   // ============================================================
   // Returns true if a certain property is set
   // ============================================================
   #LKinLang_CheckProperty := (#properties AND #propertyToCheck) = #propertyToCheck;
END_FUNCTION

FUNCTION "LKinLang_CreateParameterLookUpTable" : Void   // FC35462, SCL
TITLE = LKinLang_CreateParameterLookUpTable
{ S7_Optimized_Access := 'TRUE' }
AUTHOR : tech.team.motioncontrol@siemens.com
FAMILY : LKinLang
VERSION : 1.1
// The FC creates the parameter look up table for later use in parser
   VAR_INPUT
      language : Int;   // language the lookUpTable should be created for
      mode : Bool;   // 0: Commands with ParameterNameNo 1: Commands without ParameterNameNumber
   END_VAR
   VAR_OUTPUT
      error : Bool;   // TRUE: An error occurred during the execution of the FC
      lastIndexLookUp : DInt;   // last index in lookUpTable
   END_VAR
   VAR_IN_OUT
      parameterLookUpTable : Array[1.."LKINLANG_MAX_NUMBER_OF_PARAMETERS"] of "LKinLang_typeParameterLookUp";   // created parameterLookUpTable
      parameterDefaults : Variant;   // parameter defaults
      parameterCounter : Int;   // parameter counter
      errorString : String;   // error information (textual)
   END_VAR
   VAR_TEMP
      tempParameterIndex : Int;
      tempParameterDefinition : "LKinLang_typeParameterDefinition";
      tempCounter : Int;
      tempSeparator : Array[1.."LKINLANG_NUMBER_OF_SEPARATORS"] of Byte;
      tempMerger : Array[1.."LKINLANG_NUMBER_OF_MERGERS"] of Byte;
      tempParameterDefinitionEmpty : "LKinLang_typeParameterDefinition";
      tempFollowValueCounter : Int;
      tempValidCounts : "LKinLang_typePathDataElementCounter";
      tempString : "LKinLang_typeVariableDeclaration";
      tempKeyToken : "LKinLang_typeKeyToken";
   END_VAR
BEGIN
   //==========================================================================================
   // SIEMENS AG
   // (c)Copyright 2019 All Rights Reserved
   //------------------------------------------------------------------------------------------
   // Library: LKinLang
   // Tested with: S7-1517T-3 PN/DP
   // Engineering: TIA Portal V15
   // Restrictions: ---
   // Requirements: S7-1500T FW 2.5
   // Functionality: LKinLang_CreateParameterLookUpTable
   // The FC creates the parameter look up table for later use in parser
   // 
   // Support: tech.team.motioncontrol@siemens.com
   // Note: Parameter comments are only available in language 'English (United States)'
   //------------------------------------------------------------------------------------------
   // Change log table:
   // Version    Date          Expert in charge    Changes applied
   // 01.00.00   28.05.2019    FR                  First created version
   // 01.00.02   29.07.2019    FR                  Mode now part of internal IF condition
   //===========================================================================================


   //======================================================================
   // Is token a known parameter - return: parameter number for array
   //======================================================================
   // Initialize
   #tempCounter := 0;
   #tempParameterIndex := 0;

   // Check for vallid parameters
   WHILE #tempParameterIndex <> -1 DO
     "LKinLang_SelectLangPackage"(language := #language,
                                  variableDeclarations=>#tempString,
                                  keyToken=>#tempKeyToken,
                                  parameterDefinition := #tempParameterDefinition,
                                  separators => #tempSeparator,
                                  mergers => #tempMerger,
                                  validCounts => #tempValidCounts,
                                  parameterNumber := #tempParameterIndex,
                                  parameterDefaults := #parameterDefaults);


     IF (#tempParameterIndex > -1 AND #tempParameterDefinition.parameterNameNumber <> -1 AND #mode = 0) // Check parameters with parameter number (>-1)
       OR (#tempParameterIndex > -1 AND #tempParameterDefinition.parameterNameNumber = -1 AND #mode = 1) // Check parameters without parameter number (=-1)
     THEN
       #parameterLookUpTable[#parameterCounter].parameterNameString := #tempParameterDefinition.parameterNameString;
       #parameterLookUpTable[#parameterCounter].parameterNameNumber := #tempParameterDefinition.parameterNameNumber;
       #parameterLookUpTable[#parameterCounter].parameterNumber := #tempParameterIndex;

       IF #tempParameterDefinition.priorities <> #tempParameterDefinitionEmpty.priorities THEN
         #parameterLookUpTable[#parameterCounter].directValueWord.%X0 := true;
       END_IF;

       IF #tempParameterDefinition.priorities.cmdCoordinates <> #tempParameterDefinitionEmpty.priorities.cmdCoordinates THEN
         #parameterLookUpTable[#parameterCounter].directValueWord.%X1 := true;
       END_IF;

       IF #tempParameterDefinition.priorities.cmdParameters <> #tempParameterDefinitionEmpty.priorities.cmdParameters THEN
         #parameterLookUpTable[#parameterCounter].directValueWord.%X2 := true;
       END_IF;
       IF #tempParameterDefinition.priorities.cmdParameters.pathDynamics <> #tempParameterDefinitionEmpty.priorities.cmdParameters.pathDynamics THEN
         #parameterLookUpTable[#parameterCounter].directValueWord.%X3 := true;
       END_IF;
       IF #tempParameterDefinition.priorities.cmdParameters.circleParameters <> #tempParameterDefinitionEmpty.priorities.cmdParameters.circleParameters THEN
         #parameterLookUpTable[#parameterCounter].directValueWord.%X4 := true;
       END_IF;

       FOR #tempFollowValueCounter := 1 TO "LKINLANG_NUMBER_OF_FOLLOW_VALUES" DO
         IF #tempParameterDefinition.followingValues[#tempFollowValueCounter] <> #tempParameterDefinitionEmpty.followingValues[#tempFollowValueCounter] THEN
           #parameterLookUpTable[#parameterCounter].followValueWords[#tempFollowValueCounter].%X0 := TRUE;
         END_IF;

         IF #tempParameterDefinition.followingValues[#tempFollowValueCounter].cmdCoordinates <> #tempParameterDefinitionEmpty.followingValues[#tempFollowValueCounter].cmdCoordinates THEN
           #parameterLookUpTable[#parameterCounter].followValueWords[#tempFollowValueCounter].%X1 := TRUE;
         END_IF;

         IF #tempParameterDefinition.followingValues[#tempFollowValueCounter].cmdParameters <> #tempParameterDefinitionEmpty.followingValues[#tempFollowValueCounter].cmdParameters THEN
           #parameterLookUpTable[#parameterCounter].followValueWords[#tempFollowValueCounter].%X2 := TRUE;
         END_IF;

         IF #tempParameterDefinition.followingValues[#tempFollowValueCounter].cmdParameters.pathDynamics <> #tempParameterDefinitionEmpty.followingValues[#tempFollowValueCounter].cmdParameters.pathDynamics THEN
           #parameterLookUpTable[#parameterCounter].followValueWords[#tempFollowValueCounter].%X3 := TRUE;
         END_IF;

         IF #tempParameterDefinition.followingValues[#tempFollowValueCounter].cmdParameters.circleParameters <> #tempParameterDefinitionEmpty.followingValues[#tempFollowValueCounter].cmdParameters.circleParameters THEN
           #parameterLookUpTable[#parameterCounter].followValueWords[#tempFollowValueCounter].%X4 := TRUE;
         END_IF;
       END_FOR;

       #parameterCounter += 1;
       #lastIndexLookUp := #parameterCounter;

       // Check ParameterCounter for Overflow
       IF #parameterCounter > "LKINLANG_MAX_NUMBER_OF_PARAMETERS" THEN
         #error := TRUE;
         #errorString := CONCAT(IN1 := #errorString, IN2 := 'Error: Array overflow lookUp table; Increase "LKINLANG_MAX_NUMBER_OF_PARAMETERS"');
         RETURN;
       END_IF;

     ELSE
       ;// no match
     END_IF;

     #tempCounter += 1;

     // Abort searching when tempParameterIndex = -1
     IF #tempParameterIndex <> -1 THEN
       #tempParameterIndex := #tempCounter;
     END_IF;

   END_WHILE;
END_FUNCTION

FUNCTION "LKinLang_DeleteComment" : Void   // FC35463, SCL
TITLE = LKinLang_DeleteComment
{ S7_Optimized_Access := 'TRUE' }
AUTHOR : tech.team.motioncontrol@siemens.com
FAMILY : LKinLang
VERSION : 1.1
// The FC deletes comments from a given string
   VAR_IN_OUT
      codeline : String;   // line to edit by deleting comments
   END_VAR
   VAR_TEMP
      tempPosOfCommentSign : Int;   // temporary variable for position of found comments
   END_VAR
BEGIN
   //==========================================================================================
   // SIEMENS AG
   // (c)Copyright 2019 All Rights Reserved
   //------------------------------------------------------------------------------------------
   // Library: LKinLang
   // Tested with: S7-1517T-3 PN/DP
   // Engineering: TIA Portal V15
   // Restrictions: ---
   // Requirements: S7-1500T FW 2.5
   // Functionality: LKinLang_DeleteComment
   // The FC deletes comments from a given string
   // 
   // Support: tech.team.motioncontrol@siemens.com
   // Note: Parameter comments are only available in language 'English (United States)'
   //------------------------------------------------------------------------------------------
   // Change log table:
   // Version    Date          Expert in charge    Changes applied
   // 01.00.00   28.05.2019    FR                  First created version
   //===========================================================================================

   //======================================================================
   // Delete comment in referenced ascii line
   //======================================================================  

   // Search semicolon
   #tempPosOfCommentSign := FIND(IN1 := #codeline, IN2 := ';');
   // Get line without comment
   IF #tempPosOfCommentSign <> 0 THEN
     #codeline := MID(IN := #codeline, L := #tempPosOfCommentSign - 1, P := 1);
   END_IF;
END_FUNCTION

FUNCTION "LKinLang_DeleteMoreThanOneSpaceInRow" : Void   // FC35464, SCL
TITLE = LKinLang_DeleteMoreThanOneSpaceInRow
{ S7_Optimized_Access := 'TRUE' }
AUTHOR : tech.team.motioncontrol@siemens.com
FAMILY : LKinLang
VERSION : 1.1
// The FC deletes spaces if there are more than one in a row
   VAR_IN_OUT
      codeLine : String;   // line to edit by deleting multiple spaces
   END_VAR
   VAR_TEMP
      tempCodeLine : String["LKINLANG_LENGTH_OF_ASCII_LINE_STRING"];   // temporary variable to store string
      tempSignCounter : Int;   // temporary variable to count signs
      tempSpaceCounter : Int;   // temporary variable to count spaces
      tempStringLength : Int;   // temporary variable to store string length
      tempSpaceIndex : Int;   // temporary variable to store space index
   END_VAR
   VAR CONSTANT
      SPACE : Byte := 16#20;   // space identifier in ascii code
   END_VAR
BEGIN
   //==========================================================================================
   // SIEMENS AG
   // (c)Copyright 2019 All Rights Reserved
   //------------------------------------------------------------------------------------------
   // Library: LKinLang
   // Tested with: S7-1517T-3 PN/DP
   // Engineering: TIA Portal V15
   // Restrictions: ---
   // Requirements: S7-1500T FW 2.5
   // Functionality: LKinLang_DeleteComment
   // The FC deletes spaces if there are more than one in a row
   // 
   // Support: tech.team.motioncontrol@siemens.com
   // Note: Parameter comments are only available in language 'English (United States)'
   //------------------------------------------------------------------------------------------
   // Change log table:
   // Version    Date          Expert in charge    Changes applied
   // 01.00.00   28.05.2019    FR                  First created version
   //===========================================================================================

   //======================================================================
   // Delete more than one spaces
   //====================================================================== 

   // First delete all spaces on start and end
   // -----------------------------------------------------
   // Count spaces on start ---
   #tempSignCounter := 1;

   WHILE #codeLine[#tempSignCounter] = #SPACE DO
     #tempSignCounter := #tempSignCounter + 1;
   END_WHILE;

   // Spaces
   #codeLine := RIGHT(IN := #codeLine,
                      L := LEN(#codeLine) - (#tempSignCounter - 1));


   // Count spaces on end --- 
   #tempSignCounter := LEN(#codeLine);
   WHILE #codeLine[#tempSignCounter] = #SPACE DO
     #tempSpaceCounter := #tempSpaceCounter + 1;
     #tempSignCounter := #tempSignCounter - 1;
   END_WHILE;

   #codeLine := LEFT(IN := #codeLine,
                     L := LEN(#codeLine) - #tempSpaceCounter);
   #tempSpaceCounter := 0;
   // -----------------------------------------------------

   (* // Too slow FR 2019.03.13
   // Delete more than one space in the middle
   // Testing new approach FR
   // 
   #tempSpaceIndex := FIND(IN1 := #codeLine, IN2 := '  ');

   WHILE #tempSpaceIndex <> 0 DO
     #codeLine := DELETE(IN := #codeLine, L := 1, P := #tempSpaceIndex);
     #tempSpaceIndex := FIND(IN1 := #codeLine, IN2 := '  ');
   END_WHILE;

   #codeLine := #codeLine;*)


    // Check if double space is somewhere in the codeline FR 2019.03.12
   IF FIND(IN1 := #codeLine, IN2 := '  ') <> 0 THEN
     // Delete more than one space in the middle
     #tempStringLength := LEN(#codeLine);

     FOR #tempSignCounter := 1 TO (#tempStringLength) DO
       // First character
       IF #tempSignCounter = 1 AND
         #codeLine[#tempSignCounter] <> #SPACE
       THEN
         #tempCodeLine[#tempSignCounter] := #codeLine[#tempSignCounter];

         // Last character                
       ELSIF #tempSignCounter = #tempStringLength AND
         #codeLine[#tempSignCounter] <> #SPACE
       THEN
         #tempCodeLine[#tempSignCounter - #tempSpaceCounter] := #codeLine[#tempSignCounter];

         // Between first and last character
       ELSIF #tempSignCounter > 1 AND #tempSignCounter < #tempStringLength
       THEN
         // More than one spaces in a row?
         IF #codeLine[#tempSignCounter] = #SPACE AND #codeLine[#tempSignCounter + 1] = #SPACE
         THEN
           // Increment space counter
           #tempSpaceCounter := #tempSpaceCounter + 1;
         ELSE
           // Only one Space
           #tempCodeLine[#tempSignCounter - #tempSpaceCounter] := #codeLine[#tempSignCounter];
         END_IF;

         // Increment space counter if the first or last character is a space 
       ELSE
         #tempSpaceCounter := #tempSpaceCounter + 1;
       END_IF;
     END_FOR;

     // set processed code line to in_out parameter
     #codeLine := #tempCodeLine;

   ELSE
     ;// Do nothing - already finished
     //#codeLine := #codeLine;
   END_IF;
END_FUNCTION

FUNCTION "LKinLang_IsTokenMath" : Bool   // FC35465, SCL
TITLE = LKinLang_IsTokenMath
{ S7_Optimized_Access := 'TRUE' }
AUTHOR : tech.team.motioncontrol@siemens.com
FAMILY : LKinLang
VERSION : 1.1
// Checks if a token is a math expression
   VAR_INPUT
      token : String;   // Token to check
   END_VAR
   // Ret_Val : TRUE: Token is math expression; FALSE: Token is not a math expression
BEGIN
   //==========================================================================================
   // SIEMENS AG
   // (c)Copyright 2019 All Rights Reserved
   //------------------------------------------------------------------------------------------
   // Library: LKinLang
   // Tested with: S7-1517T-3 PN/DP
   // Engineering: TIA Portal V15
   // Restrictions: ---
   // Requirements: S7-1500T FW 2.5
   // Functionality: LKinLang_IsTokenMath
   // The FC checks if a given token is a math expression
   // 
   // Support: tech.team.motioncontrol@siemens.com
   // Note: Parameter comments are only available in language 'English (United States)'
   //------------------------------------------------------------------------------------------
   // Change log table:
   // Version    Date          Expert in charge    Changes applied
   // 01.00.00   17.07.2019    FR                  First created version
   //===========================================================================================

   // Check if token is a valid math expression
   IF #token = 'SIN'
     OR #token = 'COS'  
     OR #token = 'SQR'
     OR #token = 'SQRT'
     OR #token = 'sin'
     OR #token = 'cos'
     OR #token = 'sqr'
     OR #token = 'sqrt'
   THEN
     #LKinLang_IsTokenMath := TRUE; // return true if regular math expression
   ELSE
     #LKinLang_IsTokenMath := FALSE; // return false if not
   END_IF;
END_FUNCTION

FUNCTION "LKinLang_GetValue" : DWord   // FC35466, SCL
TITLE = LKinLang_GetValue
{ S7_Optimized_Access := 'TRUE' }
AUTHOR : tech.team.motioncontrol@siemens.com
FAMILY : LKinLang
VERSION : 1.1
// The FC gets the numerical value of a given string expression
   VAR_INPUT
      tokenNo : Int;   // token number to get the numerical value for
      properties : DWord;   // properties to be considered
      followValCounter : Int;   // counter for follow value
   END_VAR
   VAR_OUTPUT
      parameterValue : LReal;   // numerical value of the expression
   END_VAR
   VAR_IN_OUT
      stringExpression : String;   // string to be checked
      errorString : String;   // error information (textual)
      token : "LKinLang_typeLineTokens";   // token information
   END_VAR
   VAR_TEMP
      tempSeparatorFound : Bool;   // temporary variable for found / not found separator
      tempStringExpression : String;   // temporary variable for storage of string expression
      tempStringLength : Int;   // temporary variable for string length
      tempCounter : Int;   // temporary counter variable
      tempSeparatorCounter : Int;   // temporary counter variable for separators
      tempTokenOffset : Int;   // temporary variable for offset of token
      tempMathParserResult : Struct   // temporary variable for math parser result
         finalResult : LReal;
         errorID : DInt;
      END_STRUCT;
   END_VAR
   VAR CONSTANT
      REAL_MIN : LReal := -3.402823E+38;
      REAL_MAX : LReal := 3.402823E+38;
      DINT_MIN : DInt := -2147483648;
      DINT_MAX : DInt := +2147483647;
      INT_MIN : Int := -32768;
      INT_MAX : Int := 32767;
      ERR_PARAMETER_COUNTER : DWord := 16#8001;
      ERR_SYNTAX_MATH_EXPRESSION : DWord := 16#8002;
      ERR_SYNTAX_PARAMETER : DWord := 16#8003;
      ERR_PARAMETER_OVERFLOW : DWord := 16#8004;
      ERR_ALREADY_SET : DWord := 16#8005;
      WARN_NO_MORE_VALUES : DWord := 16#7100;
      COMMA : Char := ',';
   END_VAR
BEGIN
   //==========================================================================================
   // SIEMENS AG
   // (c)Copyright 2019 All Rights Reserved
   //------------------------------------------------------------------------------------------
   // Library: LKinLang
   // Tested with: S7-1517T-3 PN/DP
   // Engineering: TIA Portal V15
   // Restrictions: ---
   // Requirements: S7-1500T FW 2.5
   // Functionality: LKinLang_GetValue
   // The FC gets the numerical value of a given string expression
   // 
   // Support: tech.team.motioncontrol@siemens.com
   // Note: Parameter comments are only available in language 'English (United States)'
   //------------------------------------------------------------------------------------------
   // Change log table:
   // Version    Date          Expert in charge    Changes applied
   // 01.00.00   28.05.2019    FR                  First created version
   // 01.00.01   16.01.2020    FR                  Updated to work with H functions
   //===========================================================================================

   // Initialize variables
   #LKinLang_GetValue := 0;
   #parameterValue := 0;

   // Check if the string expression contains a function separator (COMMA in this case)
   // If true copy only the string expression until the separator and leave the rest (and delete the first separator)
   #tempStringLength := LEN(#stringExpression);

   // Check for comma in stringExpression
   FOR #tempCounter := 1 TO #tempStringLength DO
     // Search for separator 
     IF #stringExpression[#tempCounter] = #COMMA THEN
       #tempSeparatorFound := TRUE;
       EXIT;
     ELSE
       #tempSeparatorFound := FALSE;
     END_IF;
   END_FOR;

   // Check if comma was found
   IF #tempSeparatorFound THEN
     // Copy first value to TempStringExpression 
     #tempStringExpression := LEFT(IN := #stringExpression, L := #tempCounter - 1);
     // Delete first from stringExpression
     #stringExpression := RIGHT(IN := #stringExpression, L := #tempStringLength - #tempCounter);
   ELSE
     #tempStringExpression := #stringExpression;
     #stringExpression := '';
   END_IF;

   IF #tempStringExpression = '' THEN
     // Empty String --> no more Values follow
     // #Lxxx_GetValue := #ERR_SYNTAX_PARAMETER;
     // #errorString := CONCAT(IN1 := #errorString, IN2 := ';Error: Missing assignment'); // Line number is added outside
     // #errorString := CONCAT(IN1 := #errorString, IN2 := INT_TO_STRING(#followValCounter)); // Line number is added outside
     RETURN;
   ELSIF #tempStringExpression = '*' THEN
     // Do not set this value
     RETURN;
   END_IF;

   IF #followValCounter > 1 THEN
     #tempSeparatorCounter := 1;
     // Check for line token offset
     FOR #tempCounter := #tokenNo TO 1 BY -1 DO
       IF #token.lineToken[#tempCounter] = #COMMA OR #token.lineToken[#tempCounter]= '=' THEN
         #tempSeparatorCounter += 1;
       END_IF;

       IF #tempSeparatorCounter = #followValCounter THEN
         EXIT;
       END_IF;
     END_FOR;
     #tempTokenOffset := #tokenNo - #tempCounter;
   ELSE
     #tempCounter := 0;
     #tempTokenOffset := 0;
   END_IF;

   // Calc LReal value --> Check Equation
   REGION GET_VALUE
     IF "LKinLang_CheckProperty"(properties := #properties, propertyToCheck := "LKINLANG_EQUATION") THEN
       REGION EQUATION
         // Equation is possible
         // 
         // Check for correct syntax
         // Two possibilities:
         // 1. Only a number after Parameter 
         // --> Equal sign is optional 
         //  --> When no equal sign then no spaces are allowed --> Example: X12
         //  --> When equal sign then one space allowed --> Example: X = 12
         // 2. Expression after Parameter
         // --> Equal sign is mandatory
         //  --> No spaces --> Example: X=12+34
         //  --> One space allowed --> Example: X = 12+34
         // 
         IF "LKinLang_PostEqualsSignWhenExpressionMandCnd"(currentTokenNo := #tokenNo,
                                                             stringExpression := #tempStringExpression,
                                                             tokenOffset := #tempTokenOffset,
                                                             lineToken := #token) 
         THEN
           // Number: just convert string to real
           IF "LKinLang_IsTokenNumberInclSign"(#tempStringExpression) THEN
             // Set parameter
             #parameterValue := STRING_TO_LREAL(#tempStringExpression);
           ELSE
             //FR not necessary //#errorString := CONCAT(IN1 := #errorString, IN2 := CONCAT(IN1 := ';Error: str=', IN2 := #tempStringExpression));
             #tempMathParserResult := "LKinLang_CalcMathAndBool"(inputString := #tempStringExpression);

             // Error with math parser
             //******************************************
             IF #tempMathParserResult.errorID <> 0 THEN
               #LKinLang_GetValue := #ERR_SYNTAX_MATH_EXPRESSION;

               #errorString := CONCAT(IN1 := #errorString, IN2 := CONCAT(IN1 := ';Error: Mathresult=', IN2 := "LKinLang_LRealToReducedString"(input:=#tempMathParserResult.finalResult,decimalPlaces:=4)));
               #errorString := CONCAT(IN1 := #errorString, IN2 := CONCAT(IN1 := ';Error: No=', IN2 := DINT_TO_STRING(#tempMathParserResult.errorID)));
               // Line number is added outside
               //#errorString := CONCAT(IN1 := #errorString, IN2 := DINT_TO_STRING(#token.lineNo));
               RETURN;
               // Math parser delivers a valid result
               //******************************************
             ELSE
               // Set parameter
               #parameterValue := #tempMathParserResult.finalResult;
             END_IF;
           END_IF;
           #tempStringExpression := '';
         ELSE
           // SyntaxError: not "Y =" or "Y19"
           #LKinLang_GetValue := #ERR_SYNTAX_PARAMETER;
           #errorString := CONCAT(IN1 := #errorString, IN2 := ';Error: Incorrect assignment (Y= or Y1)'); // Line number is added outside
           RETURN;
         END_IF;
       END_REGION EQUATION

     ELSE

       REGION NO_EQUATION
         // Equation is not possible
         IF "LKinLang_PostNumberMandCnd"(algebraicSignAllowed := True, currentTokenNo := #tokenNo, tokenOffset := #tempTokenOffset, lineTokens := #token)
         THEN
           IF "LKinLang_IsTokenNumber"(#tempStringExpression) THEN
             IF #followValCounter = 1 THEN
               #parameterValue := STRING_TO_LREAL(#token.lineToken[#tokenNo - 1]);
             ELSE
               #parameterValue := STRING_TO_LREAL(#token.lineToken[#tokenNo - #tempTokenOffset - 1]);
             END_IF;

             // Check if Mxx stands alone, also there could be something like this Mxx=29
             IF STRING_TO_LREAL(#tempStringExpression) = #parameterValue THEN
               #tempStringExpression := '';
             ELSE
               #LKinLang_GetValue := #ERR_SYNTAX_PARAMETER;
               #errorString := CONCAT(IN1 := #errorString, IN2 := ';Error: Incorrect assignment '); // Line number is added outside
               #errorString := CONCAT(IN1 := #errorString, IN2 := INT_TO_STRING(#followValCounter)); // Line number is added outside
               RETURN;
             END_IF;

           ELSIF "LKinLang_IsTokenNumberInclSign"(#tempStringExpression) THEN

             IF #followValCounter = 1 THEN
               #parameterValue := STRING_TO_LREAL(CONCAT(IN1 := #token.lineToken[#tokenNo - 1], IN2 := #token.lineToken[#tokenNo - 2]));
             ELSE
               #parameterValue := STRING_TO_LREAL(CONCAT(IN1 := #token.lineToken[#tokenNo - #tempTokenOffset - 1], IN2 := #token.lineToken[#tokenNo - #tempTokenOffset - 2]));
             END_IF;

             // Check if Mxx stands alone, also there could be something like this Mxx=29
             IF STRING_TO_LREAL(#tempStringExpression) = #parameterValue THEN
               #tempStringExpression := '';
             ELSE
               #LKinLang_GetValue := #ERR_SYNTAX_PARAMETER;
               #errorString := CONCAT(IN1 := #errorString, IN2 := ';Error: Incorrect assignment '); // Line number is added outside
               #errorString := CONCAT(IN1 := #errorString, IN2 := INT_TO_STRING(#followValCounter)); // Line number is added outside
               RETURN;
             END_IF;
           END_IF;
         ELSE
           // SyntaxError: no number after parameter
           #LKinLang_GetValue := #ERR_SYNTAX_PARAMETER;
           #errorString := CONCAT(IN1 := #errorString, IN2 := ';Error: No number after parameter'); // Line number is added outside
           RETURN;
         END_IF;
       END_REGION NO_EQUATION

     END_IF;

   END_REGION GET_VALUE
END_FUNCTION

FUNCTION "LKinLang_EvaluateCondition" : Bool   // FC35467, SCL
TITLE = LKinLang_EvaluateCondition
{ S7_Optimized_Access := 'TRUE' }
AUTHOR : tech.team.motioncontrol@siemens.com
FAMILY : LKinLang
VERSION : 1.0
// Evaluate a given condition for conditional jumps etc.
   VAR_INPUT
      offsetLastTokenIndex : UInt;   // Number of token to skip from end
   END_VAR
   VAR_IN_OUT
      tokenizedLine : "LKinLang_typeLineTokens";   // Actual tokenized line
      varRefList : "LKinLang_typeVarRefList";   // Variables reference list
      localVariables : "LKinLang_typeLocalVariables";   // Local variables array
      interfaceVariables : "LKinLang_typeInterfaceVariables";   // Interface varaibles array
      keyToken : "LKinLang_typeKeyToken";   // Key token to find variables
      subPrgList : "LKinLang_typeSubPrgList";
      errorString : String;   // error string connection
   END_VAR
   VAR_TEMP
      tempStateIntern : Int;   // Internal state
      tempTokenCounter : Int;   // Temporary counter for token
      tempVarType : Int;   // Variable type
      tempVarIndex : Int;   // Variable index in reference list
      tempStringExpression : String;   // Stringexpression
      tempTokenCheck : Struct   // Struct with the token to check / Static struct with the token to check
         actual : String;
         previous : String;
      END_STRUCT;
      tempMathParserResult : "LKinLang_typeMathParserResult";   // Result of math and bool calculation
   END_VAR
   // Ret_Val : Returns result of condition
   VAR CONSTANT
      STATE_IS_TOKEN_VARIABLE : Int := 250;   // Internal FB state: Is token variable
      STATE_TOKEN_IS_VARIABLE : Int := 260;   // Internal FB state: Token is variable
      STATE_TOKEN_IS_UNKNOWN : Int := 270;   // Internal FB state: Token is unknown
      STATE_ERROR : Int := 900;   // Internal FB state: Error
   END_VAR
BEGIN
   //==========================================================================================
   // SIEMENS AG
   // (c)Copyright 2020 All Rights Reserved
   //------------------------------------------------------------------------------------------
   // Library: LKinLang
   // Tested with: S7-1517T-3 PN/DP
   // Engineering: TIA Portal V15
   // Restrictions: ---
   // Requirements: S7-1500T FW 2.5
   // Functionality: LKinLang_EvaluateCondition
   // The FC creates a valid expression for MathParser and returns the result of the calculation
   // 
   // Support: tech.team.motioncontrol@siemens.com
   // Note: Parameter comments are only available in language 'English (United States)'
   //------------------------------------------------------------------------------------------
   // Change log table:
   // Version    Date          Expert in charge    Changes applied
   // 01.00.00   09.01.2019    FR                  First created version
   // 01.00.01   24.11.2020    FR                  Use functions to check if token is a variable
   //===========================================================================================
   //
   // Add everything except " " to the string expression 
   // If it is a variable then replace with the value of the variable
   // Call MathParser to get result of condition

   // There is no left side of equation as the "=" in a condition is not used as a assignment

   // Iterate over all token
   FOR #tempTokenCounter := 1 TO #tokenizedLine.numberOfToken - #offsetLastTokenIndex DO

     // Init variables for each loop
     #tempTokenCheck.actual := #tokenizedLine.lineToken[#tempTokenCounter];

     //Get previous token
     IF #tempTokenCounter > 1 THEN
       #tempTokenCheck.previous := #tokenizedLine.lineToken[#tempTokenCounter - 1];
     ELSE
       #tempTokenCheck.previous := '';
     END_IF;

     // Next state: IS_TOKEN_VARIABLE
     #tempStateIntern := #STATE_IS_TOKEN_VARIABLE;

     // ------------------------------------------------------------------------------------------
     // Is token variable
     // Check if token is a defined variable or interface variable
     // YES: Go to TOKEN_IS_VARIABLE
     // NO: Go to TOKEN_IS_UNKNOWN
     // ------------------------------------------------------------------------------------------ 
     REGION IS_TOKEN_VARIABLE
       IF #tempStateIntern = #STATE_IS_TOKEN_VARIABLE THEN
         // Check if token is a local or interface variable 
         "LKinLang_IsTokenVariable"(lineNumber := #tokenizedLine.lineNo,
                                    tokenCheck := #tempTokenCheck,
                                    varIndex => #tempVarIndex,
                                    varType => #tempVarType,
                                    varRefList := #varRefList,
                                    keyToken := #keyToken,
                                    subPrgList:=#subPrgList,
                                    errorString := #errorString,
                                    stringExpression := #tempStringExpression);

         // Decide where to go next
         IF #errorString <> '' THEN
           // Error occured
           #tempStateIntern := #STATE_ERROR;
           EXIT;
         ELSIF #tempVarIndex <> 0 OR #tempVarType <> 0 THEN
           // Go to "TOKEN_IS_VARIABLE"
           #tempStateIntern := #STATE_TOKEN_IS_VARIABLE;
         ELSE
           // Go to "TOKEN_IS_UNKNOWN"
           #tempStateIntern := #STATE_TOKEN_IS_UNKNOWN;
         END_IF;
       END_IF;
     END_REGION IS_TOKEN_VARIABLE

     // ------------------------------------------------------------------------------------------
     // Token is a variable
     // Token was found to be a valid variable
     // SET or GET value of variable depending on context
     // ------------------------------------------------------------------------------------------ 
     REGION TOKEN_IS_VARIABLE
       IF #tempStateIntern = #STATE_TOKEN_IS_VARIABLE THEN
         // Token is variable 
         // Decide if value of variable has to be set or value must be read
         "LKinLang_GetVariable"(varIndex:=#tempVarIndex,
                                varType:=#tempVarType,
                                localVariables:=#localVariables,
                                interfaceVariables:=#interfaceVariables,
                                stringExpression:=#tempStringExpression);
       END_IF;
     END_REGION TOKEN_IS_VARIABLE

     // ------------------------------------------------------------------------------------------
     // Token is unknown
     // Token is not a parameter or a separator 
     // Check if equation is active and add token to string expression 
     // If token consists of letters, it is a unknown parameter and a error is thrown
     // Always go to TOKEN_PROCESSED
     // ------------------------------------------------------------------------------------------ 
     REGION TOKEN_IS_UNKNOWN
       IF #tempStateIntern = #STATE_TOKEN_IS_UNKNOWN
       THEN
         // Check if actual token is not space --> Copy to StringExpression (e.g. math expressions)
         IF #tempTokenCheck.actual = 'TRUE' THEN
           #tempStringExpression := CONCAT(IN1 := '1', IN2 := #tempStringExpression);
         ELSIF #tempTokenCheck.actual = 'FALSE' THEN
           #tempStringExpression := CONCAT(IN1 := '0', IN2 := #tempStringExpression);
         ELSIF  #tempTokenCheck.actual <> ' ' THEN
           #tempStringExpression := CONCAT(IN1 := #tempTokenCheck.actual, IN2 := #tempStringExpression);
         ELSE
           ; // Do not copy "space"  into string expression
         END_IF;
       END_IF;
     END_REGION TOKEN_IS_UNKNOWN
   END_FOR;

   #LKinLang_EvaluateCondition := FALSE;

   IF #tempStateIntern <> #STATE_ERROR THEN
     // All token are processed 
     // Call MathParser and calculate result
     #tempMathParserResult := "LKinLang_CalcMathAndBool"(inputString := #tempStringExpression);

     // Check for error in math parser
     IF #tempMathParserResult.errorID <> 0
       OR #tempMathParserResult.finalResult < 0
       OR #tempMathParserResult.finalResult > 1
     THEN
       #tempStateIntern := #STATE_ERROR;
       #errorString := CONCAT(IN1 := #errorString, IN2 := ';Error: Cannot evaluate condition ');
       #errorString := CONCAT(IN1 := #errorString, IN2 := #tempStringExpression);
       #errorString := CONCAT(IN1 := #errorString, IN2 := '; in line: ');
       #errorString := CONCAT(IN1 := #errorString, IN2 := UDINT_TO_STRING(#tokenizedLine.lineNo));
     ELSE
       // Math parser delivers a valid result
       // Assign result to value
       #LKinLang_EvaluateCondition := (#tempMathParserResult.finalResult = 1); // If result = 1 then true else false
     END_IF;
   ELSE
     ; // Error occured --> Do nothing
   END_IF;
END_FUNCTION

FUNCTION "LKinLang_IsNewCommand" : Bool   // FC35469, SCL
TITLE = LKinLang_IsNewCommand
{ S7_Optimized_Access := 'TRUE' }
AUTHOR : tech.team.motioncontrol@siemens.com
FAMILY : LKinLang
VERSION : 1.1
// This function checks if a parsed line results in a new PathData command
   VAR_IN_OUT
      actualPathData : "LKinLang_typePathDataElement";   // actual PathData element to be checked
      emptyPathData : "LKinLang_typePathDataElement";   // empty PathData element for comparison
      positioningMode : Int;   // mode for positioning
   END_VAR
   VAR_TEMP
      tempCircMode0 : Bool;   // temporary variable for circMode 0
      tempCircMode1 : Bool;   // temporary variable for circMode 1
      tempCircMode2 : Bool;   // temporary variable for circMode 2
   END_VAR
BEGIN
   //==========================================================================================
   // SIEMENS AG
   // (c)Copyright 2019 All Rights Reserved
   //------------------------------------------------------------------------------------------
   // Library: LKinLang
   // Tested with: S7-1517T-3 PN/DP
   // Engineering: TIA Portal V15
   // Restrictions: ---
   // Requirements: S7-1500T FW 2.5
   // Functionality: LKinLang_IsNewCommand
   // This function checks if a parsed line results in a new PathData command
   // 
   // Support: tech.team.motioncontrol@siemens.com
   // Note: Parameter comments are only available in language 'English (United States)'
   //------------------------------------------------------------------------------------------
   // Change log table:
   // Version    Date          Expert in charge    Changes applied
   // 01.00.00   28.05.2019    FR                  First created version
   // 01.00.01   10.12.2020    FR                  Added case for cmdType=-1
   //===========================================================================================

   #LKinLang_IsNewCommand := 0;

   CASE #actualPathData.pathDataElement.cmdType OF
       -1: // Only check position
           #LKinLang_IsNewCommand := (#actualPathData.priority.cmdCoordinates.cartesianPosition.x > "LKINLANG_PRIO_UNRELEVANT")
           OR (#actualPathData.priority.cmdCoordinates.cartesianPosition.y > "LKINLANG_PRIO_UNRELEVANT")
           OR (#actualPathData.priority.cmdCoordinates.cartesianPosition.z > "LKINLANG_PRIO_UNRELEVANT")
           OR (#actualPathData.priority.cmdCoordinates.cartesianPosition.a > "LKINLANG_PRIO_UNRELEVANT");


     1,2:  // Linear command
       IF #positioningMode = 1 THEN
         // Is it a new absolute position ?
         // Check if last position is same as actual ? --> Do not check could be usefull with flags on same position
         // (#actualPathData.pathDataElement.cmdCoordinates <> #oldPathData.pathDataElement.cmdCoordinates)
         // AND
         //#LKinLang_IsNewCommand := (#actualPathData.pathDataElement.cmdCoordinates.cartesianPosition <> #emptyPathData.pathDataElement.cmdCoordinates.cartesianPosition);
         #LKinLang_IsNewCommand := (#actualPathData.priority.cmdCoordinates.cartesianPosition.x > "LKINLANG_PRIO_UNRELEVANT")
         OR (#actualPathData.priority.cmdCoordinates.cartesianPosition.y > "LKINLANG_PRIO_UNRELEVANT")
         OR (#actualPathData.priority.cmdCoordinates.cartesianPosition.z > "LKINLANG_PRIO_UNRELEVANT")
         OR (#actualPathData.priority.cmdCoordinates.cartesianPosition.a > "LKINLANG_PRIO_UNRELEVANT");

       ELSIF #positioningMode = 2 THEN
         // Is it a new relative position ?
         //#LKinLang_IsNewCommand := (#actualPathData.pathDataElement.cmdCoordinates.cartesianPosition <> #emptyPathData.pathDataElement.cmdCoordinates.cartesianPosition);
         #LKinLang_IsNewCommand := (#actualPathData.priority.cmdCoordinates.cartesianPosition.x > "LKINLANG_PRIO_UNRELEVANT")
         OR (#actualPathData.priority.cmdCoordinates.cartesianPosition.y > "LKINLANG_PRIO_UNRELEVANT")
         OR (#actualPathData.priority.cmdCoordinates.cartesianPosition.z > "LKINLANG_PRIO_UNRELEVANT")
         OR (#actualPathData.priority.cmdCoordinates.cartesianPosition.a > "LKINLANG_PRIO_UNRELEVANT");

       ELSE
         #LKinLang_IsNewCommand := FALSE;
       END_IF;

     3,4:  // Circular command
       // Is a absolute circle set ?
       // CircMode 0 // Aux Point + End Point
       #tempCircMode0 :=
       ((#actualPathData.priority.cmdCoordinates.cartesianPosition.x > "LKINLANG_PRIO_UNRELEVANT")
       OR (#actualPathData.priority.cmdCoordinates.cartesianPosition.y > "LKINLANG_PRIO_UNRELEVANT")
       OR (#actualPathData.priority.cmdCoordinates.cartesianPosition.z > "LKINLANG_PRIO_UNRELEVANT")
       OR (#actualPathData.priority.cmdCoordinates.cartesianPosition.a > "LKINLANG_PRIO_UNRELEVANT"))
       AND
       ((#actualPathData.priority.cmdParameters.circleParameters.auxPoint[1] > "LKINLANG_PRIO_UNRELEVANT")
       OR (#actualPathData.priority.cmdParameters.circleParameters.auxPoint[2] > "LKINLANG_PRIO_UNRELEVANT")
       OR (#actualPathData.priority.cmdParameters.circleParameters.auxPoint[3] > "LKINLANG_PRIO_UNRELEVANT"));

       // CircMode 1 // Aux Point + Arc
       #tempCircMode1 :=
       (#actualPathData.priority.cmdParameters.circleParameters.arc > "LKINLANG_PRIO_UNRELEVANT")
       AND
       ((#actualPathData.priority.cmdParameters.circleParameters.auxPoint[1] > "LKINLANG_PRIO_UNRELEVANT")
       OR (#actualPathData.priority.cmdParameters.circleParameters.auxPoint[2] > "LKINLANG_PRIO_UNRELEVANT")
       OR (#actualPathData.priority.cmdParameters.circleParameters.auxPoint[3] > "LKINLANG_PRIO_UNRELEVANT"));;

       // CircMode 2 // Radius + End Point
       #tempCircMode2 :=
       #actualPathData.priority.cmdParameters.circleParameters.radius > "LKINLANG_PRIO_UNRELEVANT"
       AND
       ((#actualPathData.priority.cmdCoordinates.cartesianPosition.x > "LKINLANG_PRIO_UNRELEVANT")
       OR (#actualPathData.priority.cmdCoordinates.cartesianPosition.y > "LKINLANG_PRIO_UNRELEVANT")
       OR (#actualPathData.priority.cmdCoordinates.cartesianPosition.z > "LKINLANG_PRIO_UNRELEVANT")
       OR (#actualPathData.priority.cmdCoordinates.cartesianPosition.a > "LKINLANG_PRIO_UNRELEVANT"));


       #LKinLang_IsNewCommand := #tempCircMode0 OR #tempCircMode1 OR #tempCircMode2;

     40: // Tool off
       #LKinLang_IsNewCommand := TRUE;

     41: // Tool left
       #LKinLang_IsNewCommand := TRUE;

     42: // Tool right
       #LKinLang_IsNewCommand := TRUE;

     100: // Wait time
       #LKinLang_IsNewCommand := TRUE;
     ELSE  // Statement section ELSE
       ;
   END_CASE;
END_FUNCTION

FUNCTION "LKinLang_IsTokenNumber" : Bool   // FC35470, SCL
TITLE = LKinLang_IsTokenNumber
{ S7_Optimized_Access := 'TRUE' }
AUTHOR : tech.team.motioncontrol@siemens.com
FAMILY : LKinLang
VERSION : 1.1
// The FC checks if a given token is a number
   VAR_INPUT
      tokenToCheck : String[254];   // token to be checked
   END_VAR
   VAR_TEMP
      tempSignIndex : Int;   // temporary variable storing the index sign
   END_VAR
   // Ret_Val : TRUE: token is number; FALSE: token is NOT a number
BEGIN
   //==========================================================================================
   // SIEMENS AG
   // (c)Copyright 2019 All Rights Reserved
   //------------------------------------------------------------------------------------------
   // Library: LKinLang
   // Tested with: S7-1517T-3 PN/DP
   // Engineering: TIA Portal V15
   // Restrictions: ---
   // Requirements: S7-1500T FW 2.5
   // Functionality: LKinLang_IsTokenNumber
   // The FC checks if a given token is a number
   // 
   // Support: tech.team.motioncontrol@siemens.com
   // Note: Parameter comments are only available in language 'English (United States)'
   //------------------------------------------------------------------------------------------
   // Change log table:
   // Version    Date          Expert in charge    Changes applied
   // 01.00.00   28.05.2019    FR                  First created version
   //===========================================================================================

   //======================================================================
   // Is token (or any other string) a number - return: yes or no
   //======================================================================
   // Initialize temp variables
   #tempSignIndex := 0;

   // Initialize --> no match
   #LKinLang_IsTokenNumber := TRUE;
   // Check for all valid parameters
   FOR #tempSignIndex := 1 TO LEN(#tokenToCheck) DO
     // Match?
     IF NOT "LKinLang_CharacterIsNumeric"(#tokenToCheck[#tempSignIndex]) THEN
       #LKinLang_IsTokenNumber := FALSE;
       EXIT;
     ELSE
       ;// no match
     END_IF;
   END_FOR;
END_FUNCTION

FUNCTION "LKinLang_IsTokenNumberInclSign" : Bool   // FC35471, SCL
TITLE = LKinLang_IsTokenNumberInclSign
{ S7_Optimized_Access := 'TRUE' }
AUTHOR : tech.team.motioncontrol@siemens.com
FAMILY : LKinLang
VERSION : 1.1
// The FC checks if a given token is a number including a sign
   VAR_INPUT
      tokenToCheck : String;   // token to be checked
   END_VAR
   VAR_TEMP
      tempSignIndex : Int;   // temporary variable storing the index sign
   END_VAR
   // Ret_Val : TRUE: token is including a sign;FALSE: token is NOT including a sign
BEGIN
   //==========================================================================================
   // SIEMENS AG
   // (c)Copyright 2019 All Rights Reserved
   //------------------------------------------------------------------------------------------
   // Library: LKinLang
   // Tested with: S7-1517T-3 PN/DP
   // Engineering: TIA Portal V15
   // Restrictions: ---
   // Requirements: S7-1500T FW 2.5
   // Functionality: LKinLang_IsTokenNumberInclSign
   // The FC checks if a given token is a number including a sign
   // 
   // Support: tech.team.motioncontrol@siemens.com
   // Note: Parameter comments are only available in language 'English (United States)'
   //------------------------------------------------------------------------------------------
   // Change log table:
   // Version    Date          Expert in charge    Changes applied
   // 01.00.00   28.05.2019    FR                  First created version
   //===========================================================================================

   //======================================================================
   // Is token (or any other string) a number  OR a number inlcusive algebraic sign
   // Return: yes or no
   //======================================================================

   #tempSignIndex :=0;

   // Initialize --> no match
   #LKinLang_IsTokenNumberInclSign := TRUE;
   // Check for all valid parameters
   FOR #tempSignIndex := 1 TO LEN(#tokenToCheck) DO
     // Match?
     IF "LKinLang_CharacterIsNumeric"(#tokenToCheck[#tempSignIndex])
       // Check for algebraic sign
       OR (#tempSignIndex = 1 AND (#tokenToCheck[1] = '+' OR #tokenToCheck[1] = '-'))
     THEN
       ; // match

     ELSE // no match
       #LKinLang_IsTokenNumberInclSign := FALSE;
       EXIT;
     END_IF;
   END_FOR;
END_FUNCTION

FUNCTION "LKinLang_IsTokenParameter" : USInt   // FC35472, SCL
TITLE = LKinLang_IsTokenParameter
{ S7_Optimized_Access := 'TRUE' }
AUTHOR : tech.team.motioncontrol@siemens.com
FAMILY : LKinLang